DATA_BLOCK "PN_FlowRate"   // DB1003
{ S7_Optimized_Access := 'FALSE' }
VERSION : 0.1
   VAR
      SetIndex : Int := 1;
      ActIndex : Int := 1;
      Send : Bool := FALSE;
      IndexError : Bool := FALSE;   // Maximaler Index wurde überschritten
      Component : Array[0..16] of Struct
         FlowC : "IDM_402_Analogout_Flow_Controller";   // FlowC
         Flow_F : "IDM_115_FlowSpeedFloat";   // Flow
         FlowC_F : "IDM_415_Analogout_Flow_Controller_Float";
      END_STRUCT;
   END_VAR
BEGIN
   Component[1].FlowC_F.Address := 1000;
   Component[2].FlowC_F.Address := 1100;
   Component[2].FlowC_F.Active := TRUE;
   Component[1].FlowC_F.Active := TRUE;
   Component[0].FlowC.Address := 16#0000;
   Component[0].FlowC.Active := FALSE;
   Component[0].FlowC.ChckConnFault := FALSE;
   Component[0].FlowC.ChckConnDone := FALSE;
   Component[0].FlowC.GeneralParameters.Request := FALSE;
   Component[0].FlowC.GeneralParameters.Transmitting := FALSE;
   Component[0].FlowC.GeneralParameters.Active := FALSE;
   Component[0].FlowC.GeneralParameters.Data.Kalibrierfaktor := 10000;
   Component[0].FlowC.GeneralParameters.Data.MaxDurchfluss := 1000;
   Component[0].FlowC.GeneralParameters.Data.Nachstellzeit := 50;
   Component[0].FlowC.GeneralParameters.Data.Filterzeit := 200;
   Component[0].FlowC.Grenzen.Request := FALSE;
   Component[0].FlowC.Grenzen.Transmitting := FALSE;
   Component[0].FlowC.Grenzen.Active := FALSE;
   Component[0].FlowC.Grenzen.Data.ObergrenzeStellgröße := 10000;
   Component[0].FlowC.Grenzen.Data.UntergrenzeStellgröße := 0;
   Component[0].FlowC.Grenzen.Data.VerzögerungAlarmObergrenze := 1000;
   Component[0].FlowC.Grenzen.Data.VerzögerungAlarmUntergrenze := 1000;
   Component[0].FlowC.SkalierungAI.Request := FALSE;
   Component[0].FlowC.SkalierungAI.Transmitting := FALSE;
   Component[0].FlowC.SkalierungAI.Active := FALSE;
   Component[0].FlowC.SkalierungAI.Data.Bereichsobergrenze := 10000;
   Component[0].FlowC.SkalierungAI.Data.Bereichsuntergrenze := -10000;
   Component[0].FlowC.SkalierungAI.Data.Mittelwertzeit := 100;
   Component[0].Flow_F.Address := 0;
   Component[0].Flow_F.Active := FALSE;
   Component[0].Flow_F.ChckConnFault := FALSE;
   Component[0].Flow_F.ChckConnDone := FALSE;
   Component[0].Flow_F.Skalierung.Request := FALSE;
   Component[0].Flow_F.Skalierung.Transmitting := FALSE;
   Component[0].Flow_F.Skalierung.Active := FALSE;
   Component[0].Flow_F.Skalierung.Data.Kalibrierfaktor := 0.0;
   Component[0].Flow_F.Skalierung.Data.Filterzeit := 16#0000;
   Component[0].FlowC_F.Address := 1000;
   Component[0].FlowC_F.Active := TRUE;
   Component[0].FlowC_F.ChckConnFault := FALSE;
   Component[0].FlowC_F.ChckConnDone := FALSE;
   Component[0].FlowC_F."I/O".InputData.Flow := 0.0;
   Component[0].FlowC_F."I/O".InputData.Weight := 0.0;
   Component[0].FlowC_F."I/O".InputData.ActPresSDA := 0;
   Component[0].FlowC_F."I/O".InputData.Control.ZeroFlow := FALSE;
   Component[0].FlowC_F."I/O".InputData.Control.SDAactiv := FALSE;
   Component[0].FlowC_F."I/O".InputData.Control.FlowControlUpperLimit := FALSE;
   Component[0].FlowC_F."I/O".InputData.Control.FlowControlLowerLimit := FALSE;
   Component[0].FlowC_F."I/O".InputData.Control.FlowLowerLimit := FALSE;
   Component[0].FlowC_F."I/O".InputData.Control.FlowUpperLimit := FALSE;
   Component[0].FlowC_F."I/O".InputData.Control.Spare06 := FALSE;
   Component[0].FlowC_F."I/O".InputData.Control.Spare07 := FALSE;
   Component[0].FlowC_F."I/O".OutputData.Flow := 0.0;
   Component[0].FlowC_F."I/O".OutputData.FlowSDA := 0.0;
   Component[0].FlowC_F."I/O".OutputData.PressSDA := 0.0;
   Component[0].FlowC_F."I/O".OutputData.actPressSDA := 0.0;
   Component[0].FlowC_F."I/O".OutputData.Control.NonControledValue := FALSE;
   Component[0].FlowC_F."I/O".OutputData.Control.ControledValue := FALSE;
   Component[0].FlowC_F."I/O".OutputData.Control.SetValueOverlay := FALSE;
   Component[0].FlowC_F."I/O".OutputData.Control.SDATrig := FALSE;
   Component[0].FlowC_F."I/O".OutputData.Control.ResetWeight := FALSE;
   Component[0].FlowC_F."I/O".OutputData.Control.Spare05 := FALSE;
   Component[0].FlowC_F."I/O".OutputData.Control.Spare06 := FALSE;
   Component[0].FlowC_F."I/O".OutputData.Control.Spare07 := FALSE;
   Component[0].FlowC_F.Hardware.Request := TRUE;
   Component[0].FlowC_F.Hardware.Transmitting := FALSE;
   Component[0].FlowC_F.Hardware.Active := FALSE;
   Component[0].FlowC_F.Hardware.Data.AO_Ausgangskanal_FU := 16#00;
   Component[0].FlowC_F.Hardware.Data.AI_Eingangskanal_Druck := 16#00;
   Component[0].FlowC_F.Hardware.Data.DI_Eingangskanal_Puls := 16#00;
   Component[0].FlowC_F.Hardware.Data.Konfig1 := 16#41;
   Component[0].FlowC_F.Hardware.Data.Konfig2 := 16#00;
   Component[0].FlowC_F.Hardware.Data.Rampenzeit := 0.1;
   Component[0].FlowC_F.GeneralParameters.Request := TRUE;
   Component[0].FlowC_F.GeneralParameters.Transmitting := FALSE;
   Component[0].FlowC_F.GeneralParameters.Active := FALSE;
   Component[0].FlowC_F.GeneralParameters.Data.Kalibrierfaktor := 3.165003;
   Component[0].FlowC_F.GeneralParameters.Data.MaxDurchfluss := 703.3333;
   Component[0].FlowC_F.GeneralParameters.Data.Nachstellzeit := 0.3;
   Component[0].FlowC_F.GeneralParameters.Data.Filterzeit := 0.2;
   Component[0].FlowC_F.Grenzen.Request := TRUE;
   Component[0].FlowC_F.Grenzen.Tranmitting := FALSE;
   Component[0].FlowC_F.Grenzen.Active := FALSE;
   Component[0].FlowC_F.Grenzen.Data.ObergrenzeStellgröße := 1.0;
   Component[0].FlowC_F.Grenzen.Data.UntergrenzeStellgröße := 0.0;
   Component[0].FlowC_F.Grenzen.Data.VerzögerungAlarmObergrenze := 1.0;
   Component[0].FlowC_F.Grenzen.Data.VerzögerungAlarmUntergrenze := 2.0;
   Component[0].FlowC_F.SkalierungAI.Request := TRUE;
   Component[0].FlowC_F.SkalierungAI.Transmitting := FALSE;
   Component[0].FlowC_F.SkalierungAI.Data.Bereichsobergrenze := 600.0;
   Component[0].FlowC_F.SkalierungAI.Data.Bereichsuntergrenze := 0.0;
   Component[0].FlowC_F.SkalierungAI.Data.Mittelwertzeit := 0.1;
   Component[0].FlowC_F.Visualisierung.BetriebsartAnalogausgang := 16#01;
   Component[0].FlowC_F.Visualisierung.BipolarerAusgang := 16#00;
   Component[0].FlowC_F.Visualisierung.Polarität := 16#00;
   Component[0].FlowC_F.Visualisierung.BetriebsartAnalogeingang := 16#02;
   Component[0].FlowC_F.Visualisierung.BetriebsartQuadraturdekoder := 16#00;
   Component[0].FlowC_F.Visualisierung.QuelleIstdruck := 16#00;
   Component[0].FlowC_F.Visualisierung.Dichte := 0.0;
   Component[1].FlowC.Address := 16#0000;
   Component[1].FlowC.Active := FALSE;
   Component[1].FlowC.ChckConnFault := FALSE;
   Component[1].FlowC.ChckConnDone := FALSE;
   Component[1].FlowC.GeneralParameters.Request := FALSE;
   Component[1].FlowC.GeneralParameters.Transmitting := FALSE;
   Component[1].FlowC.GeneralParameters.Active := FALSE;
   Component[1].FlowC.GeneralParameters.Data.Kalibrierfaktor := 10000;
   Component[1].FlowC.GeneralParameters.Data.MaxDurchfluss := 1000;
   Component[1].FlowC.GeneralParameters.Data.Nachstellzeit := 50;
   Component[1].FlowC.GeneralParameters.Data.Filterzeit := 200;
   Component[1].FlowC.Grenzen.Request := FALSE;
   Component[1].FlowC.Grenzen.Transmitting := FALSE;
   Component[1].FlowC.Grenzen.Active := FALSE;
   Component[1].FlowC.Grenzen.Data.ObergrenzeStellgröße := 10000;
   Component[1].FlowC.Grenzen.Data.UntergrenzeStellgröße := 0;
   Component[1].FlowC.Grenzen.Data.VerzögerungAlarmObergrenze := 1000;
   Component[1].FlowC.Grenzen.Data.VerzögerungAlarmUntergrenze := 1000;
   Component[1].FlowC.SkalierungAI.Request := FALSE;
   Component[1].FlowC.SkalierungAI.Transmitting := FALSE;
   Component[1].FlowC.SkalierungAI.Active := FALSE;
   Component[1].FlowC.SkalierungAI.Data.Bereichsobergrenze := 10000;
   Component[1].FlowC.SkalierungAI.Data.Bereichsuntergrenze := -10000;
   Component[1].FlowC.SkalierungAI.Data.Mittelwertzeit := 100;
   Component[1].Flow_F.Address := 0;
   Component[1].Flow_F.Active := FALSE;
   Component[1].Flow_F.ChckConnFault := FALSE;
   Component[1].Flow_F.ChckConnDone := FALSE;
   Component[1].Flow_F.Skalierung.Request := FALSE;
   Component[1].Flow_F.Skalierung.Transmitting := FALSE;
   Component[1].Flow_F.Skalierung.Active := FALSE;
   Component[1].Flow_F.Skalierung.Data.Kalibrierfaktor := 0.0;
   Component[1].Flow_F.Skalierung.Data.Filterzeit := 16#0000;
   Component[1].FlowC_F.ChckConnFault := FALSE;
   Component[1].FlowC_F.ChckConnDone := FALSE;
   Component[1].FlowC_F."I/O".InputData.Flow := 0.0;
   Component[1].FlowC_F."I/O".InputData.Weight := 0.0;
   Component[1].FlowC_F."I/O".InputData.ActPresSDA := 0;
   Component[1].FlowC_F."I/O".InputData.Control.ZeroFlow := FALSE;
   Component[1].FlowC_F."I/O".InputData.Control.SDAactiv := FALSE;
   Component[1].FlowC_F."I/O".InputData.Control.FlowControlUpperLimit := FALSE;
   Component[1].FlowC_F."I/O".InputData.Control.FlowControlLowerLimit := FALSE;
   Component[1].FlowC_F."I/O".InputData.Control.FlowLowerLimit := FALSE;
   Component[1].FlowC_F."I/O".InputData.Control.FlowUpperLimit := FALSE;
   Component[1].FlowC_F."I/O".InputData.Control.Spare06 := FALSE;
   Component[1].FlowC_F."I/O".InputData.Control.Spare07 := FALSE;
   Component[1].FlowC_F."I/O".OutputData.Flow := 0.0;
   Component[1].FlowC_F."I/O".OutputData.FlowSDA := 0.0;
   Component[1].FlowC_F."I/O".OutputData.PressSDA := 0.0;
   Component[1].FlowC_F."I/O".OutputData.actPressSDA := 0.0;
   Component[1].FlowC_F."I/O".OutputData.Control.NonControledValue := FALSE;
   Component[1].FlowC_F."I/O".OutputData.Control.ControledValue := FALSE;
   Component[1].FlowC_F."I/O".OutputData.Control.SetValueOverlay := FALSE;
   Component[1].FlowC_F."I/O".OutputData.Control.SDATrig := FALSE;
   Component[1].FlowC_F."I/O".OutputData.Control.ResetWeight := FALSE;
   Component[1].FlowC_F."I/O".OutputData.Control.Spare05 := FALSE;
   Component[1].FlowC_F."I/O".OutputData.Control.Spare06 := FALSE;
   Component[1].FlowC_F."I/O".OutputData.Control.Spare07 := FALSE;
   Component[1].FlowC_F.Hardware.Request := TRUE;
   Component[1].FlowC_F.Hardware.Transmitting := FALSE;
   Component[1].FlowC_F.Hardware.Active := FALSE;
   Component[1].FlowC_F.Hardware.Data.AO_Ausgangskanal_FU := 16#00;
   Component[1].FlowC_F.Hardware.Data.AI_Eingangskanal_Druck := 16#00;
   Component[1].FlowC_F.Hardware.Data.DI_Eingangskanal_Puls := 16#00;
   Component[1].FlowC_F.Hardware.Data.Konfig1 := 16#41;
   Component[1].FlowC_F.Hardware.Data.Konfig2 := 16#00;
   Component[1].FlowC_F.Hardware.Data.Rampenzeit := 0.1;
   Component[1].FlowC_F.GeneralParameters.Request := FALSE;
   Component[1].FlowC_F.GeneralParameters.Transmitting := FALSE;
   Component[1].FlowC_F.GeneralParameters.Active := FALSE;
   Component[1].FlowC_F.GeneralParameters.Data.Kalibrierfaktor := 3.165003;
   Component[1].FlowC_F.GeneralParameters.Data.MaxDurchfluss := 703.3333;
   Component[1].FlowC_F.GeneralParameters.Data.Nachstellzeit := 0.3;
   Component[1].FlowC_F.GeneralParameters.Data.Filterzeit := 0.2;
   Component[1].FlowC_F.Grenzen.Request := FALSE;
   Component[1].FlowC_F.Grenzen.Tranmitting := FALSE;
   Component[1].FlowC_F.Grenzen.Active := FALSE;
   Component[1].FlowC_F.Grenzen.Data.ObergrenzeStellgröße := 1.0;
   Component[1].FlowC_F.Grenzen.Data.UntergrenzeStellgröße := 0.0;
   Component[1].FlowC_F.Grenzen.Data.VerzögerungAlarmObergrenze := 1.0;
   Component[1].FlowC_F.Grenzen.Data.VerzögerungAlarmUntergrenze := 2.0;
   Component[1].FlowC_F.SkalierungAI.Request := FALSE;
   Component[1].FlowC_F.SkalierungAI.Transmitting := FALSE;
   Component[1].FlowC_F.SkalierungAI.Data.Bereichsobergrenze := 600.0;
   Component[1].FlowC_F.SkalierungAI.Data.Bereichsuntergrenze := 0.0;
   Component[1].FlowC_F.SkalierungAI.Data.Mittelwertzeit := 0.1;
   Component[1].FlowC_F.Visualisierung.BetriebsartAnalogausgang := 16#01;
   Component[1].FlowC_F.Visualisierung.BipolarerAusgang := 16#00;
   Component[1].FlowC_F.Visualisierung.Polarität := 16#00;
   Component[1].FlowC_F.Visualisierung.BetriebsartAnalogeingang := 16#02;
   Component[1].FlowC_F.Visualisierung.BetriebsartQuadraturdekoder := 16#00;
   Component[1].FlowC_F.Visualisierung.QuelleIstdruck := 16#00;
   Component[1].FlowC_F.Visualisierung.Dichte := 0.0;
   Component[2].FlowC.Address := 16#0000;
   Component[2].FlowC.Active := FALSE;
   Component[2].FlowC.ChckConnFault := FALSE;
   Component[2].FlowC.ChckConnDone := FALSE;
   Component[2].FlowC.GeneralParameters.Request := FALSE;
   Component[2].FlowC.GeneralParameters.Transmitting := FALSE;
   Component[2].FlowC.GeneralParameters.Active := FALSE;
   Component[2].FlowC.GeneralParameters.Data.Kalibrierfaktor := 10000;
   // 1534 more start values not shown
END_DATA_BLOCK

DATA_BLOCK "PN_CON"   // DB1004
{ S7_Optimized_Access := 'FALSE' }
VERSION : 0.1
   VAR
      Dataset : "SZL-IDW#16#xy96_DataSet";
   END_VAR
BEGIN
   Dataset.LogicalAddr := 16#0000;
   Dataset.System := 16#0000;
   Dataset.API := 16#0000_0000;
   Dataset.Station := 16#0000;
   Dataset.Slot := 16#0000;
   Dataset.Subslot := 16#0000;
   Dataset.Offset := 16#0000;
   Dataset.SetType.Herstellernummer := 16#0000;
   Dataset.SetType.Geraet := 16#0000;
   Dataset.SetType.LaufendeNummer := 16#0000;
   Dataset.SetType.ModulIdentifikation1 := 16#0000;
   Dataset.SetType.ModulIdentifikation2 := 16#0000;
   Dataset.SetType.SubmodulIdentifikation1 := 16#0000;
   Dataset.SetType.Submodulidentifikation2 := 16#0000;
   Dataset.SetType_UnEqual_ActualType[0] := FALSE;
   Dataset.SetType_UnEqual_ActualType[1] := FALSE;
   Dataset.SetType_UnEqual_ActualType[2] := FALSE;
   Dataset.SetType_UnEqual_ActualType[3] := FALSE;
   Dataset.SetType_UnEqual_ActualType[4] := FALSE;
   Dataset.SetType_UnEqual_ActualType[5] := FALSE;
   Dataset.SetType_UnEqual_ActualType[6] := FALSE;
   Dataset.SetType_UnEqual_ActualType[7] := FALSE;
   Dataset.SetType_UnEqual_ActualType[8] := FALSE;
   Dataset.SetType_UnEqual_ActualType[9] := FALSE;
   Dataset.SetType_UnEqual_ActualType[10] := FALSE;
   Dataset.SetType_UnEqual_ActualType[11] := FALSE;
   Dataset.SetType_UnEqual_ActualType[12] := FALSE;
   Dataset.SetType_UnEqual_ActualType[13] := FALSE;
   Dataset.SetType_UnEqual_ActualType[14] := FALSE;
   Dataset.SetType_UnEqual_ActualType[15] := FALSE;
   Dataset.res := 16#0000;
   Dataset.IOStat.BaugruppeWartungsbedarf := FALSE;
   Dataset.IOStat.BaugruppeWartungsanforderung := FALSE;
   Dataset.IOStat.res10 := FALSE;
   Dataset.IOStat.res11 := FALSE;
   Dataset.IOStat.res12 := FALSE;
   Dataset.IOStat.res13 := FALSE;
   Dataset.IOStat.res14 := FALSE;
   Dataset.IOStat.res15 := FALSE;
   Dataset.IOStat.BaugruppeGestoert := FALSE;
   Dataset.IOStat.BaugruppeVorhanden := FALSE;
   Dataset.IOStat.BaugruppeNichtVerfuegbar := FALSE;
   Dataset.IOStat.BaugruppeDeaktiviert := FALSE;
   Dataset.IOStat.StoerungDerStation := FALSE;
   Dataset.IOStat.M7_BaugruppeHostFuerSup := FALSE;
   Dataset.IOStat.res6 := FALSE;
   Dataset.IOStat.BaugruppeImLokalbussegment := FALSE;
   Dataset.AreaID_ModuleWidth := 16#0000;
   Dataset.res_1 := 16#0000;
   Dataset.res_2 := 16#0000;
   Dataset.res_3 := 16#0000;
   Dataset.res_4 := 16#0000;
   Dataset.res_5 := 16#0000;
   Dataset.res_6 := 16#0000;
   Dataset.res_7 := 16#0000;
   Dataset.res_8 := 16#0000;
   Dataset.res_9 := 16#0000;
   Dataset.res_10 := 16#0000;
END_DATA_BLOCK

DATA_BLOCK "PN_DeviceState"   // DB1005
TITLE = ProfiNetState
{ S7_Optimized_Access := 'TRUE' }
VERSION : 0.1
   VAR
      StatePN : Array[1..1023] of Bool;
      StateModulPN : Array[1..1023] of Bool;
   END_VAR
BEGIN
   StatePN[1] := TRUE;
   StatePN[2] := TRUE;
   StatePN[3] := TRUE;
   StatePN[4] := TRUE;
   StatePN[5] := TRUE;
   StatePN[6] := TRUE;
   StatePN[7] := FALSE;
   StatePN[8] := FALSE;
   StatePN[9] := FALSE;
   StatePN[10] := FALSE;
   StatePN[11] := FALSE;
   StatePN[12] := FALSE;
   StatePN[13] := FALSE;
   StatePN[14] := FALSE;
   StatePN[15] := FALSE;
   StatePN[16] := FALSE;
   StatePN[17] := FALSE;
   StatePN[18] := FALSE;
   StatePN[19] := FALSE;
   StatePN[20] := FALSE;
   StatePN[21] := FALSE;
   StatePN[22] := FALSE;
   StatePN[23] := FALSE;
   StatePN[24] := FALSE;
   StatePN[25] := FALSE;
   StatePN[26] := FALSE;
   StatePN[27] := FALSE;
   StatePN[28] := FALSE;
   StatePN[29] := FALSE;
   StatePN[30] := FALSE;
   StatePN[31] := FALSE;
   StatePN[32] := TRUE;
   StatePN[33] := TRUE;
   StatePN[34] := FALSE;
   StatePN[35] := FALSE;
   StatePN[36] := FALSE;
   StatePN[37] := FALSE;
   StatePN[38] := FALSE;
   StatePN[39] := FALSE;
   StatePN[40] := FALSE;
   StatePN[41] := FALSE;
   StatePN[42] := FALSE;
   StatePN[43] := FALSE;
   StatePN[44] := FALSE;
   StatePN[45] := FALSE;
   StatePN[46] := FALSE;
   StatePN[47] := FALSE;
   StatePN[48] := FALSE;
   StatePN[49] := FALSE;
   StatePN[50] := FALSE;
   StatePN[51] := FALSE;
   StatePN[52] := FALSE;
   StatePN[53] := FALSE;
   StatePN[54] := FALSE;
   StatePN[55] := FALSE;
   StatePN[56] := FALSE;
   StatePN[57] := FALSE;
   StatePN[58] := FALSE;
   StatePN[59] := FALSE;
   StatePN[60] := FALSE;
   StatePN[61] := FALSE;
   StatePN[62] := FALSE;
   StatePN[63] := FALSE;
   StatePN[64] := FALSE;
   StatePN[65] := FALSE;
   StatePN[66] := FALSE;
   StatePN[67] := FALSE;
   StatePN[68] := FALSE;
   StatePN[69] := FALSE;
   StatePN[70] := FALSE;
   StatePN[71] := FALSE;
   StatePN[72] := FALSE;
   StatePN[73] := FALSE;
   StatePN[74] := FALSE;
   StatePN[75] := FALSE;
   StatePN[76] := FALSE;
   StatePN[77] := FALSE;
   StatePN[78] := FALSE;
   StatePN[79] := FALSE;
   StatePN[80] := FALSE;
   StatePN[81] := FALSE;
   StatePN[82] := FALSE;
   StatePN[83] := FALSE;
   StatePN[84] := FALSE;
   StatePN[85] := FALSE;
   StatePN[86] := FALSE;
   StatePN[87] := FALSE;
   StatePN[88] := FALSE;
   StatePN[89] := FALSE;
   StatePN[90] := FALSE;
   StatePN[91] := FALSE;
   StatePN[92] := FALSE;
   StatePN[93] := FALSE;
   StatePN[94] := FALSE;
   StatePN[95] := FALSE;
   StatePN[96] := FALSE;
   StatePN[97] := FALSE;
   StatePN[98] := FALSE;
   StatePN[99] := FALSE;
   StatePN[100] := FALSE;
   StatePN[101] := FALSE;
   StatePN[102] := FALSE;
   StatePN[103] := FALSE;
   StatePN[104] := FALSE;
   StatePN[105] := FALSE;
   StatePN[106] := FALSE;
   StatePN[107] := FALSE;
   StatePN[108] := FALSE;
   StatePN[109] := FALSE;
   StatePN[110] := FALSE;
   StatePN[111] := FALSE;
   StatePN[112] := FALSE;
   StatePN[113] := FALSE;
   StatePN[114] := FALSE;
   StatePN[115] := FALSE;
   StatePN[116] := FALSE;
   StatePN[117] := FALSE;
   StatePN[118] := FALSE;
   StatePN[119] := FALSE;
   StatePN[120] := FALSE;
   StatePN[121] := FALSE;
   StatePN[122] := FALSE;
   StatePN[123] := FALSE;
   StatePN[124] := FALSE;
   StatePN[125] := FALSE;
   StatePN[126] := FALSE;
   StatePN[127] := FALSE;
   StatePN[128] := FALSE;
   StatePN[129] := FALSE;
   StatePN[130] := FALSE;
   StatePN[131] := FALSE;
   StatePN[132] := FALSE;
   StatePN[133] := FALSE;
   StatePN[134] := FALSE;
   StatePN[135] := FALSE;
   StatePN[136] := FALSE;
   StatePN[137] := FALSE;
   StatePN[138] := FALSE;
   StatePN[139] := FALSE;
   StatePN[140] := FALSE;
   StatePN[141] := FALSE;
   StatePN[142] := FALSE;
   StatePN[143] := FALSE;
   StatePN[144] := FALSE;
   StatePN[145] := FALSE;
   StatePN[146] := FALSE;
   StatePN[147] := FALSE;
   StatePN[148] := FALSE;
   StatePN[149] := FALSE;
   StatePN[150] := FALSE;
   StatePN[151] := FALSE;
   StatePN[152] := FALSE;
   StatePN[153] := FALSE;
   StatePN[154] := FALSE;
   StatePN[155] := FALSE;
   StatePN[156] := FALSE;
   StatePN[157] := FALSE;
   StatePN[158] := FALSE;
   StatePN[159] := FALSE;
   StatePN[160] := FALSE;
   StatePN[161] := FALSE;
   StatePN[162] := FALSE;
   StatePN[163] := FALSE;
   StatePN[164] := FALSE;
   StatePN[165] := FALSE;
   StatePN[166] := FALSE;
   StatePN[167] := FALSE;
   StatePN[168] := FALSE;
   StatePN[169] := FALSE;
   StatePN[170] := FALSE;
   StatePN[171] := FALSE;
   StatePN[172] := FALSE;
   StatePN[173] := FALSE;
   StatePN[174] := FALSE;
   StatePN[175] := FALSE;
   StatePN[176] := FALSE;
   StatePN[177] := FALSE;
   StatePN[178] := FALSE;
   StatePN[179] := FALSE;
   StatePN[180] := FALSE;
   StatePN[181] := FALSE;
   StatePN[182] := FALSE;
   StatePN[183] := FALSE;
   StatePN[184] := FALSE;
   StatePN[185] := FALSE;
   StatePN[186] := FALSE;
   StatePN[187] := FALSE;
   StatePN[188] := FALSE;
   StatePN[189] := FALSE;
   StatePN[190] := FALSE;
   StatePN[191] := FALSE;
   StatePN[192] := FALSE;
   StatePN[193] := FALSE;
   StatePN[194] := FALSE;
   StatePN[195] := FALSE;
   StatePN[196] := FALSE;
   StatePN[197] := FALSE;
   StatePN[198] := FALSE;
   StatePN[199] := FALSE;
   StatePN[200] := FALSE;
   // 1846 more start values not shown
END_DATA_BLOCK

DATA_BLOCK "PN_Mixinghead"   // DB1006
{ S7_Optimized_Access := 'FALSE' }
VERSION : 0.1
   VAR
      SetIndex : Int := 1;
      ActIndex : Int := 1;
      Send : Bool := FALSE;
      IndexError : Bool := FALSE;   // Maximaler Index wurde überschritten
      Mixinghead : Array[0..16] of Struct
         Analog : "IDM_605_Mixinghead_Analog";
         Digital : "IDM_601_Mixinghead_Digital";
         ReinigungskolbenDigital : "IDM_610_CleaningPiston_Digital";
         ReinigungskolbenGeregelt : "IDM_616_CleaningPiston_Analog_Loop";
         ReinigungskolbenGesteuert : "IDM_615_CleaningPiston_Analog";
         DüseBypass : Array[1..8] of "IDM_620_Mixinghead_NozzleBypass";
         OszillierVentile : "IDM_212_Digout_Oscillation";
         Send : Bool;
      END_STRUCT;
   END_VAR
BEGIN
   Mixinghead[1].Analog.Address := 1050;
   Mixinghead[1].Digital.Address := 1050;
   Mixinghead[1].Digital.GeneralParameters.Data.EingangskanalFreigabe := 16#20;
   Mixinghead[1].Digital.Zeiten.Data.ÜberwachungszeitÖffnen := 0.5;
   Mixinghead[1].Digital.Zeiten.Data.ÜberwachungszeitSchließen := 0.5;
   Mixinghead[1].Digital.Zeiten.Data.ErlaubtePrellzeit := 0.25;
   Mixinghead[1].ReinigungskolbenDigital.GeneralParameters.Data.EingangskanalRK_Ini := 16#01;
   Mixinghead[1].ReinigungskolbenDigital.GeneralParameters.Data.AusgangRKVentil := 16#04;
   Mixinghead[2].Digital.Address := 1150;
   Mixinghead[2].ReinigungskolbenDigital.Address := 1170;
   Mixinghead[2].Digital.GeneralParameters.Data.EingangskanalFreigabe := 16#20;
   Mixinghead[2].Digital.Zeiten.Data.ÜberwachungszeitÖffnen := 0.5;
   Mixinghead[2].Digital.Zeiten.Data.ÜberwachungszeitSchließen := 0.5;
   Mixinghead[2].Digital.Zeiten.Data.ErlaubtePrellzeit := 0.01;
   Mixinghead[2].ReinigungskolbenDigital.GeneralParameters.Data.EingangskanalRK_Ini := 16#01;
   Mixinghead[2].ReinigungskolbenDigital.GeneralParameters.Data.AusgangRKVentil := 16#04;
   Mixinghead[1].Digital.Active := TRUE;
   Mixinghead[0].Analog.Address := 1050;
   Mixinghead[0].Analog.Active := FALSE;
   Mixinghead[0].Analog.ChckConnFault := FALSE;
   Mixinghead[0].Analog.ChckConnDone := FALSE;
   Mixinghead[0].Analog.Resourcen.Request := FALSE;
   Mixinghead[0].Analog.Resourcen.Transmitting := FALSE;
   Mixinghead[0].Analog.Resourcen.Active := FALSE;
   Mixinghead[0].Analog.Resourcen.Data.EingangskanalMK_Ini.Bool0 := FALSE;
   Mixinghead[0].Analog.Resourcen.Data.EingangskanalMK_Ini.Bool1 := FALSE;
   Mixinghead[0].Analog.Resourcen.Data.EingangskanalMK_Ini.Bool2 := FALSE;
   Mixinghead[0].Analog.Resourcen.Data.EingangskanalMK_Ini.Bool3 := FALSE;
   Mixinghead[0].Analog.Resourcen.Data.EingangskanalMK_Ini.Bool4 := FALSE;
   Mixinghead[0].Analog.Resourcen.Data.EingangskanalMK_Ini.Bool5 := FALSE;
   Mixinghead[0].Analog.Resourcen.Data.EingangskanalMK_Ini.Spare6 := FALSE;
   Mixinghead[0].Analog.Resourcen.Data.EingangskanalMK_Ini.Spare7 := FALSE;
   Mixinghead[0].Analog.Resourcen.Data.EingangskanalFreigabe.Bool0 := FALSE;
   Mixinghead[0].Analog.Resourcen.Data.EingangskanalFreigabe.Bool1 := FALSE;
   Mixinghead[0].Analog.Resourcen.Data.EingangskanalFreigabe.Bool2 := FALSE;
   Mixinghead[0].Analog.Resourcen.Data.EingangskanalFreigabe.Bool3 := FALSE;
   Mixinghead[0].Analog.Resourcen.Data.EingangskanalFreigabe.Bool4 := FALSE;
   Mixinghead[0].Analog.Resourcen.Data.EingangskanalFreigabe.Bool5 := FALSE;
   Mixinghead[0].Analog.Resourcen.Data.EingangskanalFreigabe.Bool6 := FALSE;
   Mixinghead[0].Analog.Resourcen.Data.EingangskanalFreigabe.Bool7 := FALSE;
   Mixinghead[0].Analog.Resourcen.Data.AnalogerAusgang.Bool0 := FALSE;
   Mixinghead[0].Analog.Resourcen.Data.AnalogerAusgang.Bool1 := FALSE;
   Mixinghead[0].Analog.Resourcen.Data.AnalogerAusgang.Bool2 := FALSE;
   Mixinghead[0].Analog.Resourcen.Data.AnalogerAusgang.Spare3 := FALSE;
   Mixinghead[0].Analog.Resourcen.Data.AnalogerAusgang.Spare4 := FALSE;
   Mixinghead[0].Analog.Resourcen.Data.AnalogerAusgang.Spare5 := FALSE;
   Mixinghead[0].Analog.Resourcen.Data.AnalogerAusgang.Spare6 := FALSE;
   Mixinghead[0].Analog.Resourcen.Data.AnalogerAusgang.Spare7 := FALSE;
   Mixinghead[0].Analog.Resourcen.Data.Betriebsart.Bool0 := FALSE;
   Mixinghead[0].Analog.Resourcen.Data.Betriebsart.Bool1 := FALSE;
   Mixinghead[0].Analog.Resourcen.Data.Betriebsart.Bool2 := FALSE;
   Mixinghead[0].Analog.Resourcen.Data.Betriebsart.Spare3 := FALSE;
   Mixinghead[0].Analog.Resourcen.Data.Betriebsart.Spare4 := FALSE;
   Mixinghead[0].Analog.Resourcen.Data.Betriebsart.Spare5 := FALSE;
   Mixinghead[0].Analog.Resourcen.Data.Betriebsart.Spare6 := FALSE;
   Mixinghead[0].Analog.Resourcen.Data.Betriebsart.Spare7 := FALSE;
   Mixinghead[0].Analog.Resourcen.Data.MischkopfKanal.Bool0 := FALSE;
   Mixinghead[0].Analog.Resourcen.Data.MischkopfKanal.Bool1 := FALSE;
   Mixinghead[0].Analog.Resourcen.Data.MischkopfKanal.Spare2 := FALSE;
   Mixinghead[0].Analog.Resourcen.Data.MischkopfKanal.Spare3 := FALSE;
   Mixinghead[0].Analog.Resourcen.Data.MischkopfKanal.Spare4 := FALSE;
   Mixinghead[0].Analog.Resourcen.Data.MischkopfKanal.Spare5 := FALSE;
   Mixinghead[0].Analog.Resourcen.Data.MischkopfKanal.Spare6 := FALSE;
   Mixinghead[0].Analog.Resourcen.Data.MischkopfKanal.Spare7 := FALSE;
   Mixinghead[0].Analog.Zeiten.Request := FALSE;
   Mixinghead[0].Analog.Zeiten.Transmitting := FALSE;
   Mixinghead[0].Analog.Zeiten.Active := FALSE;
   Mixinghead[0].Analog.Zeiten.Data.ÜberwachungszeitÖffnen := 500;
   Mixinghead[0].Analog.Zeiten.Data.ÜberwachungszeitSchließen := 500;
   Mixinghead[0].Analog.Zeiten.Data.ErlaubtePrellzeit := 20;
   Mixinghead[0].Analog.Skalierung.Request := FALSE;
   Mixinghead[0].Analog.Skalierung.Transmitting := FALSE;
   Mixinghead[0].Analog.Skalierung.Active := FALSE;
   Mixinghead[0].Analog.Skalierung.Data.Bereichsobergrenze := 10000;
   Mixinghead[0].Analog.Skalierung.Data.Bereichsuntergrenze := -10000;
   Mixinghead[0].Analog.StufenAktivierung.Request := FALSE;
   Mixinghead[0].Analog.StufenAktivierung.Transmitting := FALSE;
   Mixinghead[0].Analog.StufenAktivierung.Active := FALSE;
   Mixinghead[0].Analog.StufenAktivierung.Data.DauerStufe1 := 10;
   Mixinghead[0].Analog.StufenAktivierung.Data.DauerStufe2 := 10;
   Mixinghead[0].Analog.StufenAktivierung.Data.DauerStufe3 := 10;
   Mixinghead[0].Analog.StufenAktivierung.Data.DauerStufe4 := 10;
   Mixinghead[0].Analog.StufenAktivierung.Data.DauerStufe5 := 10;
   Mixinghead[0].Analog.StufenAktivierung.Data.LevelStufe1 := 10000;
   Mixinghead[0].Analog.StufenAktivierung.Data.LevelStufe2 := 5000;
   Mixinghead[0].Analog.StufenAktivierung.Data.LevelStufe3 := 1500;
   Mixinghead[0].Analog.StufenAktivierung.Data.LevelStufe4 := 500;
   Mixinghead[0].Analog.StufenAktivierung.Data.LevelStufe5 := 0;
   Mixinghead[0].Analog.StufenRückkehr.Request := FALSE;
   Mixinghead[0].Analog.StufenRückkehr.Transmitting := FALSE;
   Mixinghead[0].Analog.StufenRückkehr.Active := FALSE;
   Mixinghead[0].Analog.StufenRückkehr.Data.DauerStufe1 := 10;
   Mixinghead[0].Analog.StufenRückkehr.Data.DauerStufe2 := 10;
   Mixinghead[0].Analog.StufenRückkehr.Data.DauerStufe3 := 10;
   Mixinghead[0].Analog.StufenRückkehr.Data.DauerStufe4 := 10;
   Mixinghead[0].Analog.StufenRückkehr.Data.DauerStufe5 := 10;
   Mixinghead[0].Analog.StufenRückkehr.Data.LevelStufe1 := -10000;
   Mixinghead[0].Analog.StufenRückkehr.Data.LevelStufe2 := -5000;
   Mixinghead[0].Analog.StufenRückkehr.Data.LevelStufe3 := -1500;
   Mixinghead[0].Analog.StufenRückkehr.Data.LevelStufe4 := -500;
   Mixinghead[0].Analog.StufenRückkehr.Data.LevelStufe5 := 0;
   Mixinghead[0].Digital.Address := 1050;
   Mixinghead[0].Digital.Active := TRUE;
   Mixinghead[0].Digital.ChckConnFault := TRUE;
   Mixinghead[0].Digital.ChckConnDone := TRUE;
   Mixinghead[0].Digital.GeneralParameters.Request := TRUE;
   Mixinghead[0].Digital.GeneralParameters.Transmitting := TRUE;
   Mixinghead[0].Digital.GeneralParameters.Active := FALSE;
   Mixinghead[0].Digital.GeneralParameters.Data.EingangskanalMK_Ini := 16#00;
   Mixinghead[0].Digital.GeneralParameters.Data.EingangskanalFreigabe := 16#20;
   Mixinghead[0].Digital.GeneralParameters.Data.Ventilausgang := 16#00;
   Mixinghead[0].Digital.GeneralParameters.Data.MischkopfKanal := 16#00;
   Mixinghead[0].Digital.Zeiten.Request := TRUE;
   Mixinghead[0].Digital.Zeiten.Transmitting := TRUE;
   Mixinghead[0].Digital.Zeiten.Active := FALSE;
   Mixinghead[0].Digital.Zeiten.Data.ÜberwachungszeitÖffnen := 0.5;
   Mixinghead[0].Digital.Zeiten.Data.ÜberwachungszeitSchließen := 0.5;
   Mixinghead[0].Digital.Zeiten.Data.ErlaubtePrellzeit := 0.25;
   Mixinghead[0].Digital.Zeiten_2.Request := TRUE;
   Mixinghead[0].Digital.Zeiten_2.Transmitting := TRUE;
   Mixinghead[0].Digital.Zeiten_2.Active := FALSE;
   Mixinghead[0].Digital.Zeiten_2.Data.Verzögerungszeit_HW_Freigabe := 0.0;
   Mixinghead[0].ReinigungskolbenDigital.Address := 0;
   Mixinghead[0].ReinigungskolbenDigital.Active := FALSE;
   Mixinghead[0].ReinigungskolbenDigital.ChckConnFault := FALSE;
   Mixinghead[0].ReinigungskolbenDigital.ChckConnDone := FALSE;
   Mixinghead[0].ReinigungskolbenDigital.GeneralParameters.Request := TRUE;
   Mixinghead[0].ReinigungskolbenDigital.GeneralParameters.Transmitting := FALSE;
   Mixinghead[0].ReinigungskolbenDigital.GeneralParameters.Active := FALSE;
   Mixinghead[0].ReinigungskolbenDigital.GeneralParameters.Data.EingangskanalRK_Ini := 16#01;
   Mixinghead[0].ReinigungskolbenDigital.GeneralParameters.Data.AusgangRKVentil := 16#04;
   Mixinghead[0].ReinigungskolbenDigital.GeneralParameters.Data.MischkopfKanal := 16#00;
   Mixinghead[0].ReinigungskolbenDigital.Zeiten.Request := TRUE;
   Mixinghead[0].ReinigungskolbenDigital.Zeiten.Transmitting := FALSE;
   Mixinghead[0].ReinigungskolbenDigital.Zeiten.Active := FALSE;
   Mixinghead[0].ReinigungskolbenDigital.Zeiten.Data.ÜberwachungszeitVorfahren := 0.5;
   Mixinghead[0].ReinigungskolbenDigital.Zeiten.Data.ÜberwachungszeitRückfahren := 0.5;
   Mixinghead[0].ReinigungskolbenDigital.Zeiten.Data.ErlaubtePrellzeit := 0.02;
   Mixinghead[0].ReinigungskolbenDigital.Zeiten.Data.WartezeitVorne := 0.5;
   Mixinghead[0].ReinigungskolbenDigital.Zeiten.Data.VerzögerungNachSchuss := 0.5;
   Mixinghead[0].ReinigungskolbenGeregelt.Address := 0;
   Mixinghead[0].ReinigungskolbenGeregelt.Active := FALSE;
   Mixinghead[0].ReinigungskolbenGeregelt.ChckConnFault := FALSE;
   Mixinghead[0].ReinigungskolbenGeregelt.ChckConnDone := FALSE;
   Mixinghead[0].ReinigungskolbenGeregelt.GeneralParameters.Request := FALSE;
   Mixinghead[0].ReinigungskolbenGeregelt.GeneralParameters.Transmitting := FALSE;
   Mixinghead[0].ReinigungskolbenGeregelt.GeneralParameters.Active := FALSE;
   Mixinghead[0].ReinigungskolbenGeregelt.GeneralParameters.Data.AnalogerAusgang.Bool0 := FALSE;
   Mixinghead[0].ReinigungskolbenGeregelt.GeneralParameters.Data.AnalogerAusgang.Bool1 := FALSE;
   Mixinghead[0].ReinigungskolbenGeregelt.GeneralParameters.Data.AnalogerAusgang.Bool2 := FALSE;
   Mixinghead[0].ReinigungskolbenGeregelt.GeneralParameters.Data.AnalogerAusgang.Spare3 := FALSE;
   Mixinghead[0].ReinigungskolbenGeregelt.GeneralParameters.Data.AnalogerAusgang.Spare4 := FALSE;
   Mixinghead[0].ReinigungskolbenGeregelt.GeneralParameters.Data.AnalogerAusgang.Spare5 := FALSE;
   Mixinghead[0].ReinigungskolbenGeregelt.GeneralParameters.Data.AnalogerAusgang.Spare6 := FALSE;
   Mixinghead[0].ReinigungskolbenGeregelt.GeneralParameters.Data.AnalogerAusgang.Spare7 := FALSE;
   Mixinghead[0].ReinigungskolbenGeregelt.GeneralParameters.Data.Betriebsart.Bool0 := FALSE;
   Mixinghead[0].ReinigungskolbenGeregelt.GeneralParameters.Data.Betriebsart.Bool1 := FALSE;
   Mixinghead[0].ReinigungskolbenGeregelt.GeneralParameters.Data.Betriebsart.Bool2 := FALSE;
   Mixinghead[0].ReinigungskolbenGeregelt.GeneralParameters.Data.Betriebsart.Spare3 := FALSE;
   Mixinghead[0].ReinigungskolbenGeregelt.GeneralParameters.Data.Betriebsart.Spare4 := FALSE;
   Mixinghead[0].ReinigungskolbenGeregelt.GeneralParameters.Data.Betriebsart.Spare5 := FALSE;
   Mixinghead[0].ReinigungskolbenGeregelt.GeneralParameters.Data.Betriebsart.Spare6 := FALSE;
   Mixinghead[0].ReinigungskolbenGeregelt.GeneralParameters.Data.Betriebsart.Spare7 := FALSE;
   Mixinghead[0].ReinigungskolbenGeregelt.GeneralParameters.Data.AnalogerEingang.Bool0 := FALSE;
   Mixinghead[0].ReinigungskolbenGeregelt.GeneralParameters.Data.AnalogerEingang.Bool1 := FALSE;
   Mixinghead[0].ReinigungskolbenGeregelt.GeneralParameters.Data.AnalogerEingang.Bool2 := FALSE;
   Mixinghead[0].ReinigungskolbenGeregelt.GeneralParameters.Data.AnalogerEingang.Spare3 := FALSE;
   Mixinghead[0].ReinigungskolbenGeregelt.GeneralParameters.Data.AnalogerEingang.Spare4 := FALSE;
   Mixinghead[0].ReinigungskolbenGeregelt.GeneralParameters.Data.AnalogerEingang.Spare5 := FALSE;
   Mixinghead[0].ReinigungskolbenGeregelt.GeneralParameters.Data.AnalogerEingang.Spare6 := FALSE;
   Mixinghead[0].ReinigungskolbenGeregelt.GeneralParameters.Data.AnalogerEingang.Spare7 := FALSE;
   Mixinghead[0].ReinigungskolbenGeregelt.GeneralParameters.Data.Betriebsart_1.Bool0 := FALSE;
   Mixinghead[0].ReinigungskolbenGeregelt.GeneralParameters.Data.Betriebsart_1.Bool1 := FALSE;
   Mixinghead[0].ReinigungskolbenGeregelt.GeneralParameters.Data.Betriebsart_1.Spare2 := FALSE;
   Mixinghead[0].ReinigungskolbenGeregelt.GeneralParameters.Data.Betriebsart_1.Spare3 := FALSE;
   Mixinghead[0].ReinigungskolbenGeregelt.GeneralParameters.Data.Betriebsart_1.Spare4 := FALSE;
   Mixinghead[0].ReinigungskolbenGeregelt.GeneralParameters.Data.Betriebsart_1.Spare5 := FALSE;
   Mixinghead[0].ReinigungskolbenGeregelt.GeneralParameters.Data.Betriebsart_1.Spare6 := FALSE;
   Mixinghead[0].ReinigungskolbenGeregelt.GeneralParameters.Data.Betriebsart_1.Spare7 := FALSE;
   Mixinghead[0].ReinigungskolbenGeregelt.GeneralParameters.Data.MischkopfKanal.Bool0 := FALSE;
   Mixinghead[0].ReinigungskolbenGeregelt.GeneralParameters.Data.MischkopfKanal.Bool1 := FALSE;
   Mixinghead[0].ReinigungskolbenGeregelt.GeneralParameters.Data.MischkopfKanal.Spare2 := FALSE;
   Mixinghead[0].ReinigungskolbenGeregelt.GeneralParameters.Data.MischkopfKanal.Spare3 := FALSE;
   Mixinghead[0].ReinigungskolbenGeregelt.GeneralParameters.Data.MischkopfKanal.Spare4 := FALSE;
   Mixinghead[0].ReinigungskolbenGeregelt.GeneralParameters.Data.MischkopfKanal.Spare5 := FALSE;
   Mixinghead[0].ReinigungskolbenGeregelt.GeneralParameters.Data.MischkopfKanal.Spare6 := FALSE;
   Mixinghead[0].ReinigungskolbenGeregelt.GeneralParameters.Data.MischkopfKanal.Spare7 := FALSE;
   Mixinghead[0].ReinigungskolbenGeregelt.GeneralParameters.Data.MischkopfKanal.AnalogerAusgang.Bool0 := FALSE;
   Mixinghead[0].ReinigungskolbenGeregelt.GeneralParameters.Data.MischkopfKanal.AnalogerAusgang.Bool1 := FALSE;
   Mixinghead[0].ReinigungskolbenGeregelt.GeneralParameters.Data.MischkopfKanal.AnalogerAusgang.Bool2 := FALSE;
   Mixinghead[0].ReinigungskolbenGeregelt.GeneralParameters.Data.MischkopfKanal.AnalogerAusgang.Spare3 := FALSE;
   Mixinghead[0].ReinigungskolbenGeregelt.GeneralParameters.Data.MischkopfKanal.AnalogerAusgang.Spare4 := FALSE;
   Mixinghead[0].ReinigungskolbenGeregelt.GeneralParameters.Data.MischkopfKanal.AnalogerAusgang.Spare5 := FALSE;
   Mixinghead[0].ReinigungskolbenGeregelt.GeneralParameters.Data.MischkopfKanal.AnalogerAusgang.Spare6 := FALSE;
   Mixinghead[0].ReinigungskolbenGeregelt.GeneralParameters.Data.MischkopfKanal.AnalogerAusgang.Spare7 := FALSE;
   Mixinghead[0].ReinigungskolbenGeregelt.Zeiten.Request := FALSE;
   Mixinghead[0].ReinigungskolbenGeregelt.Zeiten.Transmitting := FALSE;
   Mixinghead[0].ReinigungskolbenGeregelt.Zeiten.Active := FALSE;
   Mixinghead[0].ReinigungskolbenGeregelt.Zeiten.Data.ÜberwachungszeitVorfahren := 500;
   Mixinghead[0].ReinigungskolbenGeregelt.Zeiten.Data.ÜberwachungszeitRückfahren := 500;
   // 7875 more start values not shown
END_DATA_BLOCK

DATA_BLOCK "PN_Error"   // DB1007
{ S7_Optimized_Access := 'FALSE' }
VERSION : 0.1
   VAR
      "Counter" : Int := 0;
      Fault : Bool := TRUE;   // Any fault depenDOng transmitting data to pronet
      MaxCounterExceeded : Bool := FALSE;   // Counter exceeded
      Transmitting : Bool := FALSE;   // Transmitting is not finished yet
      Reset : Bool := FALSE;
      Error : Array[1..10] of "TransmittingError";
      Module : Array[0..10] of Struct
         DO_1 : DWord;
         "DO" : DWord;
         AI : Array[1..8] of Int;
         AIr : Array[1..8] of Int;
         AO : Array[1..8] of Int;
      END_STRUCT;
   END_VAR
BEGIN
   Error[1].Address := 282;
   Error[1].Index := 3;
   Error[1].Length := 16;
   Error[1].State := 16#C080_A300;
   Error[2].Address := 282;
   Error[2].Index := 2;
   Error[2].Length := 16;
   Error[2].State := 16#C080_A300;
   Error[3].Address := 313;
   Error[3].Index := 2;
   Error[3].Length := 12;
   Error[3].State := 16#C080_A300;
   Error[4].Address := 313;
   Error[4].Index := 1;
   Error[4].Length := 4;
   Error[4].State := 16#C080_A300;
   Error[5].Address := 284;
   Error[5].Index := 4;
   Error[5].Length := 12;
   Error[5].State := 16#C080_A300;
   Error[6].Address := 284;
   Error[6].Index := 3;
   Error[6].Length := 16;
   Error[6].State := 16#C080_A300;
   Error[7].Address := 284;
   Error[7].Index := 2;
   Error[7].Length := 16;
   Error[7].State := 16#C080_A300;
   Error[8].Address := 282;
   Error[8].Index := 4;
   Error[8].Length := 12;
   Error[8].State := 16#C080_A300;
   Error[9].Address := 282;
   Error[9].Index := 3;
   Error[9].Length := 16;
   Error[9].State := 16#C080_A300;
   Error[10].Address := 282;
   Error[10].Index := 2;
   Error[10].Length := 16;
   Error[10].State := 16#C080_A300;
   Module[0].DO_1 := 16#0000_0000;
   Module[0]."DO" := 16#0000_0000;
   Module[0].AI[1] := 0;
   Module[0].AI[2] := 0;
   Module[0].AI[3] := 0;
   Module[0].AI[4] := 0;
   Module[0].AI[5] := 0;
   Module[0].AI[6] := 0;
   Module[0].AI[7] := 0;
   Module[0].AI[8] := 0;
   Module[0].AIr[1] := 0;
   Module[0].AIr[2] := 0;
   Module[0].AIr[3] := 0;
   Module[0].AIr[4] := 0;
   Module[0].AIr[5] := 0;
   Module[0].AIr[6] := 0;
   Module[0].AIr[7] := 0;
   Module[0].AIr[8] := 0;
   Module[0].AO[1] := 0;
   Module[0].AO[2] := 0;
   Module[0].AO[3] := 0;
   Module[0].AO[4] := 0;
   Module[0].AO[5] := 0;
   Module[0].AO[6] := 0;
   Module[0].AO[7] := 0;
   Module[0].AO[8] := 0;
   Module[1].DO_1 := 16#0000_0000;
   Module[1]."DO" := 16#0000_0000;
   Module[1].AI[1] := 0;
   Module[1].AI[2] := 0;
   Module[1].AI[3] := 0;
   Module[1].AI[4] := 0;
   Module[1].AI[5] := 0;
   Module[1].AI[6] := 0;
   Module[1].AI[7] := 0;
   Module[1].AI[8] := 0;
   Module[1].AIr[1] := 0;
   Module[1].AIr[2] := 0;
   Module[1].AIr[3] := 0;
   Module[1].AIr[4] := 0;
   Module[1].AIr[5] := 0;
   Module[1].AIr[6] := 0;
   Module[1].AIr[7] := 0;
   Module[1].AIr[8] := 0;
   Module[1].AO[1] := 0;
   Module[1].AO[2] := 0;
   Module[1].AO[3] := 0;
   Module[1].AO[4] := 0;
   Module[1].AO[5] := 0;
   Module[1].AO[6] := 0;
   Module[1].AO[7] := 0;
   Module[1].AO[8] := 0;
   Module[2].DO_1 := 16#0000_0000;
   Module[2]."DO" := 16#0000_0000;
   Module[2].AI[1] := 0;
   Module[2].AI[2] := 0;
   Module[2].AI[3] := 0;
   Module[2].AI[4] := 0;
   Module[2].AI[5] := 0;
   Module[2].AI[6] := 0;
   Module[2].AI[7] := 0;
   Module[2].AI[8] := 0;
   Module[2].AIr[1] := 0;
   Module[2].AIr[2] := 0;
   Module[2].AIr[3] := 0;
   Module[2].AIr[4] := 0;
   Module[2].AIr[5] := 0;
   Module[2].AIr[6] := 0;
   Module[2].AIr[7] := 0;
   Module[2].AIr[8] := 0;
   Module[2].AO[1] := 0;
   Module[2].AO[2] := 0;
   Module[2].AO[3] := 0;
   Module[2].AO[4] := 0;
   Module[2].AO[5] := 0;
   Module[2].AO[6] := 0;
   Module[2].AO[7] := 0;
   Module[2].AO[8] := 0;
   Module[3].DO_1 := 16#0000_0000;
   Module[3]."DO" := 16#0000_0000;
   Module[3].AI[1] := 0;
   Module[3].AI[2] := 0;
   Module[3].AI[3] := 0;
   Module[3].AI[4] := 0;
   Module[3].AI[5] := 0;
   Module[3].AI[6] := 0;
   Module[3].AI[7] := 0;
   Module[3].AI[8] := 0;
   Module[3].AIr[1] := 0;
   Module[3].AIr[2] := 0;
   Module[3].AIr[3] := 0;
   Module[3].AIr[4] := 0;
   Module[3].AIr[5] := 0;
   Module[3].AIr[6] := 0;
   Module[3].AIr[7] := 0;
   Module[3].AIr[8] := 0;
   Module[3].AO[1] := 0;
   Module[3].AO[2] := 0;
   Module[3].AO[3] := 0;
   Module[3].AO[4] := 0;
   Module[3].AO[5] := 0;
   Module[3].AO[6] := 0;
   Module[3].AO[7] := 0;
   Module[3].AO[8] := 0;
   Module[4].DO_1 := 16#0000_0000;
   Module[4]."DO" := 16#0000_0000;
   Module[4].AI[1] := 0;
   Module[4].AI[2] := 0;
   Module[4].AI[3] := 0;
   Module[4].AI[4] := 0;
   Module[4].AI[5] := 0;
   Module[4].AI[6] := 0;
   Module[4].AI[7] := 0;
   Module[4].AI[8] := 0;
   Module[4].AIr[1] := 0;
   Module[4].AIr[2] := 0;
   Module[4].AIr[3] := 0;
   Module[4].AIr[4] := 0;
   Module[4].AIr[5] := 0;
   Module[4].AIr[6] := 0;
   Module[4].AIr[7] := 0;
   Module[4].AIr[8] := 0;
   Module[4].AO[1] := 0;
   Module[4].AO[2] := 0;
   Module[4].AO[3] := 0;
   Module[4].AO[4] := 0;
   Module[4].AO[5] := 0;
   Module[4].AO[6] := 0;
   Module[4].AO[7] := 0;
   Module[4].AO[8] := 0;
   Module[5].DO_1 := 16#0000_0000;
   Module[5]."DO" := 16#0000_0000;
   Module[5].AI[1] := 0;
   Module[5].AI[2] := 0;
   Module[5].AI[3] := 0;
   Module[5].AI[4] := 0;
   Module[5].AI[5] := 0;
   Module[5].AI[6] := 0;
   Module[5].AI[7] := 0;
   Module[5].AI[8] := 0;
   Module[5].AIr[1] := 0;
   Module[5].AIr[2] := 0;
   Module[5].AIr[3] := 0;
   Module[5].AIr[4] := 0;
   Module[5].AIr[5] := 0;
   Module[5].AIr[6] := 0;
   Module[5].AIr[7] := 0;
   Module[5].AIr[8] := 0;
   Module[5].AO[1] := 0;
   Module[5].AO[2] := 0;
   Module[5].AO[3] := 0;
   Module[5].AO[4] := 0;
   Module[5].AO[5] := 0;
   Module[5].AO[6] := 0;
   Module[5].AO[7] := 0;
   Module[5].AO[8] := 0;
   Module[6].DO_1 := 16#0000_0000;
   Module[6]."DO" := 16#0000_0000;
   Module[6].AI[1] := 0;
   Module[6].AI[2] := 0;
   // 126 more start values not shown
END_DATA_BLOCK

DATA_BLOCK "PN_Get_DIAG"   // DB1009
TITLE = Diagnose Baugruppe
{ S7_Optimized_Access := 'TRUE' }
VERSION : 0.1
   VAR
      diagMODE : UInt := 1;
      LADDR : Hw_Any := 0;
      returnValue : Int := 0;
      CountDiagDetails : UInt := 0;
      Diag : DIS;
   END_VAR
BEGIN
   Diag.MaintainanceState := 16#0000_0000;
   Diag.ComponentStateDetail := 16#0000_8000;
   Diag.OwnState := 0;
   Diag.IOState := 16#0001;
   Diag.OperatingState := 0;
END_DATA_BLOCK

DATA_BLOCK "DB1010_TT_Fault"   // DB1010
{ S7_Optimized_Access := 'FALSE' }
VERSION : 0.1
   VAR
      ES : Struct   // Emergency stop information
         ControlCabinet : Bool;
         Machine : Bool;
         Handling_1 : Bool;
         Handling_2 : Bool;
         Operatingpanel : Bool;
         Spare_8 : Bool;
         Spare_007 : Bool;
         Spare_008 : Bool;
         Spare_009 : Bool;
         Spare_010 : Bool;
         Spare_011 : Bool;
         Spare_012 : Bool;
         Spare_013 : Bool;
         Spare_014 : Bool;
         Spare_015 : Bool;
         Spare_016 : Bool;
      END_STRUCT;
      AS : Struct   // Automatic stop information
         AS_Activ : Bool;   // Automatic stop still activ
         AS_WingDoor : Bool;   // Automatic stop wing door
         Spare_0_2 : Bool;
         Spare_0_3 : Bool;
         Spare_0_4 : Bool;
         Spare_0_5 : Bool;
         Spare_0_6 : Bool;
         Spare_0_7 : Bool;
         Spare_1_0 : Bool;
         Spare_1_1 : Bool;
         Spare_1_2 : Bool;
         Spare_1_3 : Bool;
         Spare_1_4 : Bool;
         Spare_1_5 : Bool;
         Spare_1_6 : Bool;
         Spare_1_7 : Bool;
      END_STRUCT;
   END_VAR
BEGIN
END_DATA_BLOCK

DATA_BLOCK "DB1011_TT_Fault"   // DB1011
{ S7_Optimized_Access := 'FALSE' }
AUTHOR : KT242
VERSION : 0.1
   VAR
      STG1_RT : Bool;   // Eine Störung der Gruppe 1 steht an Rundtisch 1
      STG2_RT : Bool;   // Eine Störung der Gruppe 2 steht an Rundtisch 1
      STG3_RT : Bool;   // Eine Störung der Gruppe 3 steht an Rundtisch 1
      Hupe_aus_RT : Bool;   // Merker für die Hupenquittierung bei allgemeinen Störungen Rundtisch 1
      Reset_FC_RT : Bool;   // Bit zum Zurücksetzen der Störungen in den einzelnen FC`s Rundtisch 1
      Reset_STGR_RT : Bool;   // Bit zum Zurücksetzen der Störungsbit im Stör- FC Rundtisch 1
      Stoerungsaend_RT : Bool;   // Sammelbit für eine neu anstehende Störung für Rundtisch 1
      FHM_Quitt_RT : Bool;   // Flankenmerker für die Quitiertasterauswahl Rundtisch 1
      FHM_NeuStoer_Grp_1 : Bool;   // Flankenmerker für eine neue Externe Störung der Grppe 1 für Rundtisch 1
      FHM_NeuStoer_Grp_2 : Bool;   // Flankenmerker für eine neue Externe Störung der Grppe 2 für Rundtisch 1
      FHM_NeuStoer_Grp_3 : Bool;   // Flankenmerker für eine neue Externe Störung der Grppe 3 für Rundtisch 1
      Reservebit_1_3 : Bool;
      Reservebit_1_4 : Bool;
      Reservebit_1_5 : Bool;
      Reservebit_1_6 : Bool;
      Reservebit_1_7 : Bool;
      FaultBits : Struct   // Bereich für die Speicherung der Störungen von Rundtisch 1
         Stoerung_001_016 : Word;   // RT Störungen Allgemein der Störungsgruppe I
         Stoerung_017_032 : Word;   // RT Störungen Allgemein der Störungsgruppe I
         Stoerung_033_048 : Word;   // RT Störungen Allgemein der Störungsgruppe II
         Stoerung_049_064 : Word;   // RT Störungen Allgemein der Störungsgruppe III
         Stoerung_065_080 : Word;   // RT Störungen Allgemein der Störungsgruppe III
         Stoerung_081_096 : Word;   // RT Störungen Allgemein der Störungsgruppe III
         Meldung_097_112 : Word;   // RT Meldungen Allgemein
         Meldung_113_128 : Word;   // RT Meldungen Allgemein
         Stoerung_S01 : Word;   // RT Störungen Segment 1
         Stoerung_S02 : Word;   // RT Störungen Segment 2
         Stoerung_S03 : Word;   // RT Störungen Segment 3
         Stoerung_S04 : Word;   // RT Störungen Segment 4
         Stoerung_S05 : Word;   // RT Störungen Segment 5
         Stoerung_S06 : Word;   // RT Störungen Segment 6
         Stoerung_S07 : Word;   // RT Störungen Segment 7
         Stoerung_S08 : Word;   // RT Störungen Segment 8
         Stoerung_S09 : Word;   // RT Störungen Segment 9
         Stoerung_S10 : Word;   // RT Störungen Segment 10
         Stoerung_S11 : Word;   // RT Störungen Segment 11
         Stoerung_S12 : Word;   // RT Störungen Segment 12
         Stoerung_S13 : Word;   // RT Störungen Segment 13
         Stoerung_S14 : Word;   // RT Störungen Segment 14
         Stoerung_S15 : Word;   // RT Störungen Segment 15
         Stoerung_S16 : Word;   // RT Störungen Segment 16
         Stoerung_S17 : Word;   // RT Störungen Segment 17
         Stoerung_S18 : Word;   // RT Störungen Segment 18
         Stoerung_S19 : Word;   // RT Störungen Segment 19
         Stoerung_S20 : Word;   // RT Störungen Segment 20
      END_STRUCT;
   END_VAR
BEGIN
END_DATA_BLOCK

DATA_BLOCK "DB1025_Service"   // DB1025
{ S7_Optimized_Access := 'TRUE' }
VERSION : 0.1
   VAR
      State : Struct
         Inputbyte : Byte := 16#8E;   // actual inputs from the selected byte
         Outputbyte : Byte := 16#00;   // actual outputs from the selected byte
         Spare : Int := 0;
         Spare_1 : Int := 0;
         Spare_2 : Int := 0;
         Spare_3 : Int := 0;
         Spare_4 : Int := 0;
         Spare_5 : Int := 0;
         Spare_6 : Int := 0;
         Spare_7 : Int := 0;
         Spare_8 : Int := 0;
         Spare_9 : Int := 0;
         Spare_10 : Int := 0;
         Spare_11 : Int := 0;
      END_STRUCT;
      Set : Struct
         Inputbyte : Word := 16#0000;   // input byte that should be displayed
         Outputbyte : Word := 16#0000;   // output byte that should be displayed
         Spare : Int := 0;
         Spare_1 : Int := 0;
         Spare_2 : Int := 0;
         Spare_3 : Int := 0;
         Spare_4 : Int := 0;
         Spare_5 : Int := 0;
         Spare_6 : Int := 0;
         Spare_7 : Int := 0;
         Spare_8 : Int := 0;
         Spare_9 : Int := 0;
         Spare_10 : Int := 0;
         Spare_11 : Int := 0;
      END_STRUCT;
      IP_address_Web : String := '10.100.100.101';
      IP_address_VNC : String := '10.100.100.181';
      PW_VNC : String := '8899';
   END_VAR
BEGIN
END_DATA_BLOCK

DATA_BLOCK "DB1030_TT_AddFaults"   // DB1030
{ S7_Optimized_Access := 'FALSE' }